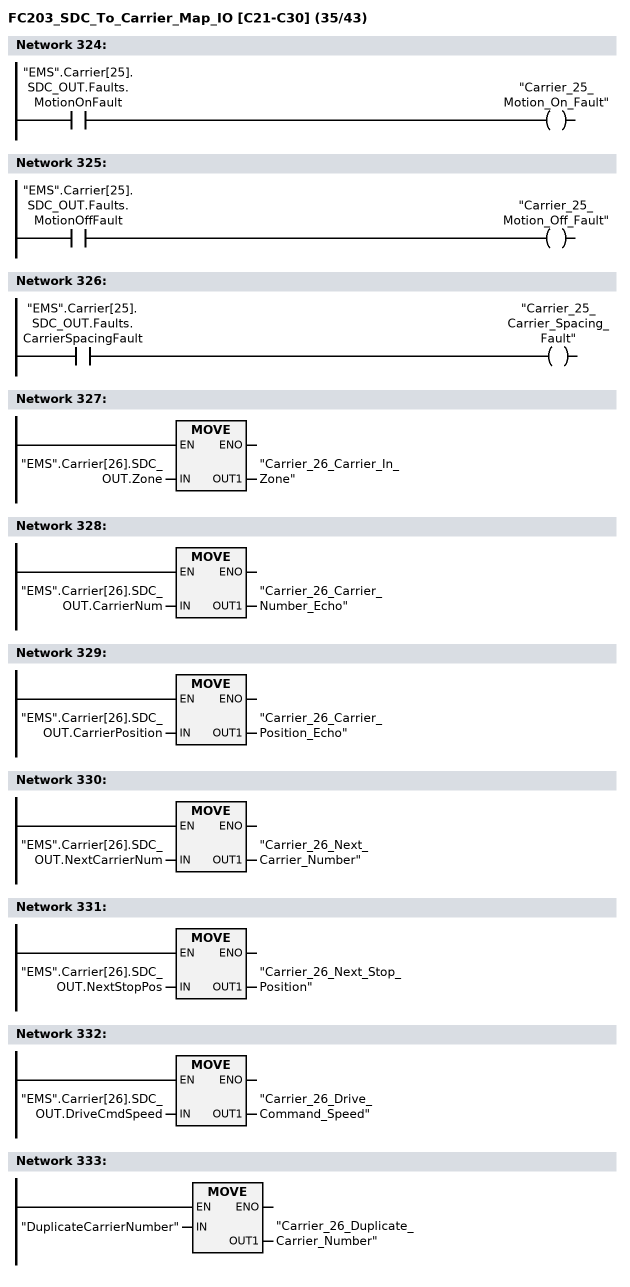
   RUNG wire#powerrail
      Contact( "EMS".Carrier[25].SDC_OUT.Faults.MotionOnFault )
      Coil( "Carrier_25_Motion_On_Fault" )
   END_RUNG
   // the same network as SCL:
   "Carrier_25_Motion_On_Fault" := "EMS".Carrier[25].SDC_OUT.Faults.MotionOnFault;
END_REGION

REGION Network 325
   RUNG wire#powerrail
      Contact( "EMS".Carrier[25].SDC_OUT.Faults.MotionOffFault )
      Coil( "Carrier_25_Motion_Off_Fault" )
   END_RUNG
   // the same network as SCL:
   "Carrier_25_Motion_Off_Fault" := "EMS".Carrier[25].SDC_OUT.Faults.MotionOffFault;
END_REGION

REGION Network 326
   RUNG wire#powerrail
      Contact( "EMS".Carrier[25].SDC_OUT.Faults.CarrierSpacingFault )
      Coil( "Carrier_25_Carrier_Spacing_Fault" )
   END_RUNG
   // the same network as SCL:
   "Carrier_25_Carrier_Spacing_Fault" := "EMS".Carrier[25].SDC_OUT.Faults.CarrierSpacingFault;
END_REGION

REGION Network 327
   RUNG wire#powerrail
      Move(in := "EMS".Carrier[26].SDC_OUT.Zone, out1 => "Carrier_26_Carrier_In_Zone")
   END_RUNG
   // the same network as SCL:
   "Carrier_26_Carrier_In_Zone" := "EMS".Carrier[26].SDC_OUT.Zone;
END_REGION

REGION Network 328
   RUNG wire#powerrail
      Move(in := "EMS".Carrier[26].SDC_OUT.CarrierNum, out1 => "Carrier_26_Carrier_Number_Echo")
   END_RUNG
   // the same network as SCL:
   "Carrier_26_Carrier_Number_Echo" := "EMS".Carrier[26].SDC_OUT.CarrierNum;
END_REGION

REGION Network 329
   RUNG wire#powerrail
      Move(in := "EMS".Carrier[26].SDC_OUT.CarrierPosition, out1 => "Carrier_26_Carrier_Position_Echo")
   END_RUNG
   // the same network as SCL:
   "Carrier_26_Carrier_Position_Echo" := "EMS".Carrier[26].SDC_OUT.CarrierPosition;
END_REGION

REGION Network 330
   RUNG wire#powerrail
      Move(in := "EMS".Carrier[26].SDC_OUT.NextCarrierNum, out1 => "Carrier_26_Next_Carrier_Number")
   END_RUNG
   // the same network as SCL:
   "Carrier_26_Next_Carrier_Number" := "EMS".Carrier[26].SDC_OUT.NextCarrierNum;
END_REGION

REGION Network 331
   RUNG wire#powerrail
      Move(in := "EMS".Carrier[26].SDC_OUT.NextStopPos, out1 => "Carrier_26_Next_Stop_Position")
   END_RUNG
   // the same network as SCL:
   "Carrier_26_Next_Stop_Position" := "EMS".Carrier[26].SDC_OUT.NextStopPos;
END_REGION

REGION Network 332
   RUNG wire#powerrail
      Move(in := "EMS".Carrier[26].SDC_OUT.DriveCmdSpeed, out1 => "Carrier_26_Drive_Command_Speed")
   END_RUNG
   // the same network as SCL:
   "Carrier_26_Drive_Command_Speed" := "EMS".Carrier[26].SDC_OUT.DriveCmdSpeed;
END_REGION

REGION Network 333
   RUNG wire#powerrail
      Move(in := "DuplicateCarrierNumber", out1 => "Carrier_26_Duplicate_Carrier_Number")
   END_RUNG
   // the same network as SCL:
   "Carrier_26_Duplicate_Carrier_Number" := "DuplicateCarrierNumber";
END_REGION

REGION Network 334
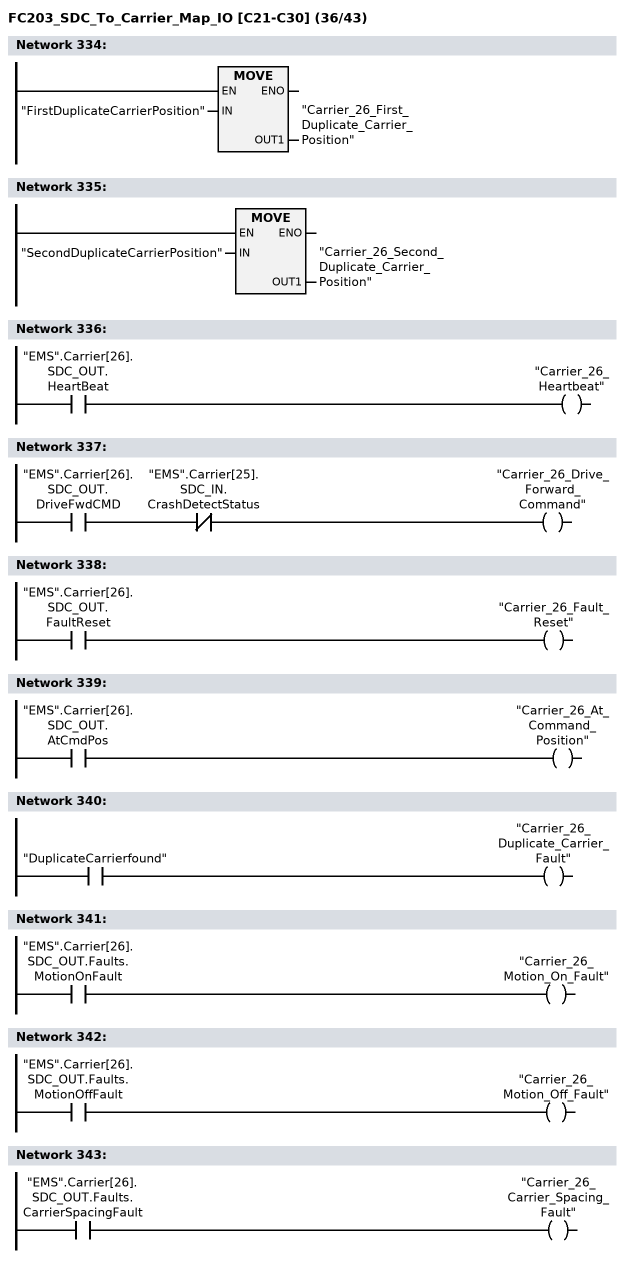
   RUNG wire#powerrail
      Move(in := "FirstDuplicateCarrierPosition", out1 => "Carrier_26_First_Duplicate_Carrier_Position")
   END_RUNG
   // the same network as SCL:
   "Carrier_26_First_Duplicate_Carrier_Position" := "FirstDuplicateCarrierPosition";
END_REGION

REGION Network 335
   RUNG wire#powerrail
      Move(in := "SecondDuplicateCarrierPosition", out1 => "Carrier_26_Second_Duplicate_Carrier_Position")
   END_RUNG
   // the same network as SCL:
   "Carrier_26_Second_Duplicate_Carrier_Position" := "SecondDuplicateCarrierPosition";
END_REGION

REGION Network 336
   RUNG wire#powerrail
      Contact( "EMS".Carrier[26].SDC_OUT.HeartBeat )
      Coil( "Carrier_26_Heartbeat" )
   END_RUNG
   // the same network as SCL:
   "Carrier_26_Heartbeat" := "EMS".Carrier[26].SDC_OUT.HeartBeat;
END_REGION

REGION Network 337
   RUNG wire#powerrail
      Contact( "EMS".Carrier[26].SDC_OUT.DriveFwdCMD )
      I_Contact( "EMS".Carrier[25].SDC_IN.CrashDetectStatus )
      Coil( "Carrier_26_Drive_Forward_Command" )
   END_RUNG
   // the same network as SCL:
   "Carrier_26_Drive_Forward_Command" := "EMS".Carrier[26].SDC_OUT.DriveFwdCMD AND NOT "EMS".Carrier[25].SDC_IN.CrashDetectStatus;
END_REGION

REGION Network 338
   RUNG wire#powerrail
      Contact( "EMS".Carrier[26].SDC_OUT.FaultReset )
      Coil( "Carrier_26_Fault_Reset" )
   END_RUNG
   // the same network as SCL:
   "Carrier_26_Fault_Reset" := "EMS".Carrier[26].SDC_OUT.FaultReset;
END_REGION

REGION Network 339
   RUNG wire#powerrail
      Contact( "EMS".Carrier[26].SDC_OUT.AtCmdPos )
      Coil( "Carrier_26_At_Command_Position" )
   END_RUNG
   // the same network as SCL:
   "Carrier_26_At_Command_Position" := "EMS".Carrier[26].SDC_OUT.AtCmdPos;
END_REGION

REGION Network 340
   RUNG wire#powerrail
      Contact( "DuplicateCarrierfound" )
      Coil( "Carrier_26_Duplicate_Carrier_Fault" )
   END_RUNG
   // the same network as SCL:
   "Carrier_26_Duplicate_Carrier_Fault" := "DuplicateCarrierfound";
END_REGION

REGION Network 341
   RUNG wire#powerrail
      Contact( "EMS".Carrier[26].SDC_OUT.Faults.MotionOnFault )
      Coil( "Carrier_26_Motion_On_Fault" )
   END_RUNG
   // the same network as SCL:
   "Carrier_26_Motion_On_Fault" := "EMS".Carrier[26].SDC_OUT.Faults.MotionOnFault;
END_REGION

REGION Network 342
   RUNG wire#powerrail
      Contact( "EMS".Carrier[26].SDC_OUT.Faults.MotionOffFault )
      Coil( "Carrier_26_Motion_Off_Fault" )
   END_RUNG
   // the same network as SCL:
   "Carrier_26_Motion_Off_Fault" := "EMS".Carrier[26].SDC_OUT.Faults.MotionOffFault;
END_REGION

REGION Network 343
   RUNG wire#powerrail
      Contact( "EMS".Carrier[26].SDC_OUT.Faults.CarrierSpacingFault )
      Coil( "Carrier_26_Carrier_Spacing_Fault" )
   END_RUNG
   // the same network as SCL:
   "Carrier_26_Carrier_Spacing_Fault" := "EMS".Carrier[26].SDC_OUT.Faults.CarrierSpacingFault;
END_REGION

REGION Network 344
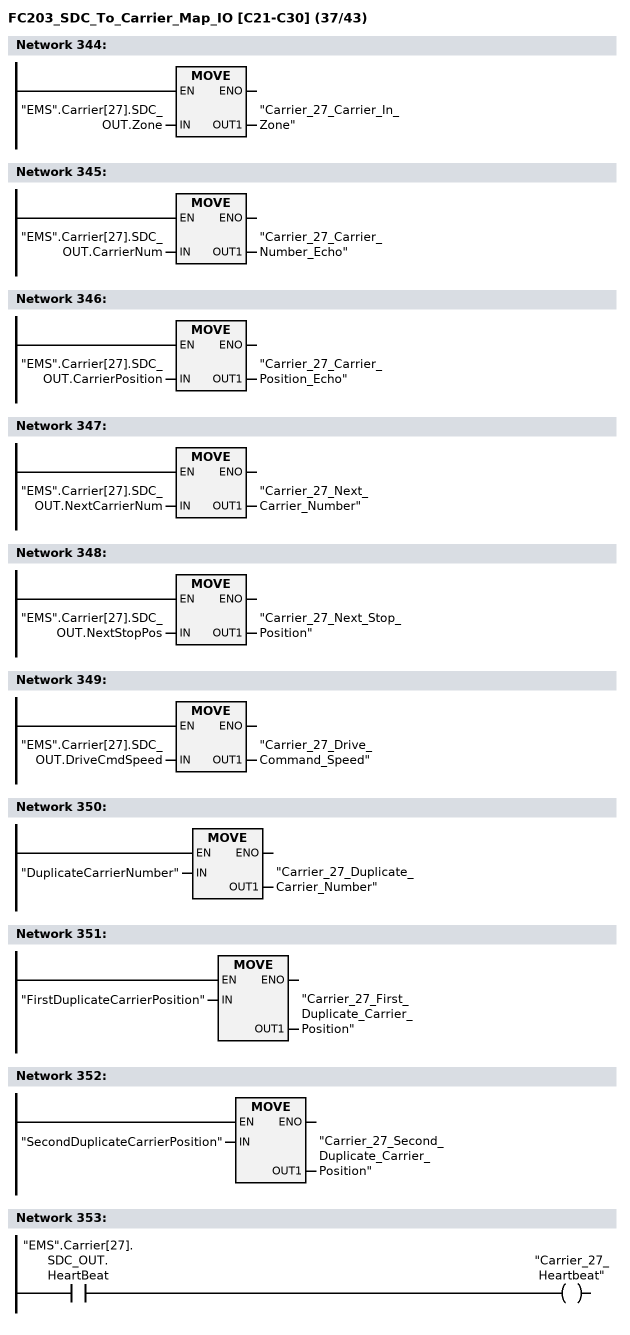
   RUNG wire#powerrail
      Move(in := "EMS".Carrier[27].SDC_OUT.Zone, out1 => "Carrier_27_Carrier_In_Zone")
   END_RUNG
   // the same network as SCL:
   "Carrier_27_Carrier_In_Zone" := "EMS".Carrier[27].SDC_OUT.Zone;
END_REGION

REGION Network 345
   RUNG wire#powerrail
      Move(in := "EMS".Carrier[27].SDC_OUT.CarrierNum, out1 => "Carrier_27_Carrier_Number_Echo")
   END_RUNG
   // the same network as SCL:
   "Carrier_27_Carrier_Number_Echo" := "EMS".Carrier[27].SDC_OUT.CarrierNum;
END_REGION

REGION Network 346
   RUNG wire#powerrail
      Move(in := "EMS".Carrier[27].SDC_OUT.CarrierPosition, out1 => "Carrier_27_Carrier_Position_Echo")
   END_RUNG
   // the same network as SCL:
   "Carrier_27_Carrier_Position_Echo" := "EMS".Carrier[27].SDC_OUT.CarrierPosition;
END_REGION

REGION Network 347
   RUNG wire#powerrail
      Move(in := "EMS".Carrier[27].SDC_OUT.NextCarrierNum, out1 => "Carrier_27_Next_Carrier_Number")
   END_RUNG
   // the same network as SCL:
   "Carrier_27_Next_Carrier_Number" := "EMS".Carrier[27].SDC_OUT.NextCarrierNum;
END_REGION

REGION Network 348
   RUNG wire#powerrail
      Move(in := "EMS".Carrier[27].SDC_OUT.NextStopPos, out1 => "Carrier_27_Next_Stop_Position")
   END_RUNG
   // the same network as SCL:
   "Carrier_27_Next_Stop_Position" := "EMS".Carrier[27].SDC_OUT.NextStopPos;
END_REGION

REGION Network 349
   RUNG wire#powerrail
      Move(in := "EMS".Carrier[27].SDC_OUT.DriveCmdSpeed, out1 => "Carrier_27_Drive_Command_Speed")
   END_RUNG
   // the same network as SCL:
   "Carrier_27_Drive_Command_Speed" := "EMS".Carrier[27].SDC_OUT.DriveCmdSpeed;
END_REGION

REGION Network 350
   RUNG wire#powerrail
      Move(in := "DuplicateCarrierNumber", out1 => "Carrier_27_Duplicate_Carrier_Number")
   END_RUNG
   // the same network as SCL:
   "Carrier_27_Duplicate_Carrier_Number" := "DuplicateCarrierNumber";
END_REGION

REGION Network 351
   RUNG wire#powerrail
      Move(in := "FirstDuplicateCarrierPosition", out1 => "Carrier_27_First_Duplicate_Carrier_Position")
   END_RUNG
   // the same network as SCL:
   "Carrier_27_First_Duplicate_Carrier_Position" := "FirstDuplicateCarrierPosition";
END_REGION

REGION Network 352
   RUNG wire#powerrail
      Move(in := "SecondDuplicateCarrierPosition", out1 => "Carrier_27_Second_Duplicate_Carrier_Position")
   END_RUNG
   // the same network as SCL:
   "Carrier_27_Second_Duplicate_Carrier_Position" := "SecondDuplicateCarrierPosition";
END_REGION

REGION Network 353
   RUNG wire#powerrail
      Contact( "EMS".Carrier[27].SDC_OUT.HeartBeat )
      Coil( "Carrier_27_Heartbeat" )
   END_RUNG
   // the same network as SCL:
   "Carrier_27_Heartbeat" := "EMS".Carrier[27].SDC_OUT.HeartBeat;
END_REGION

REGION Network 354
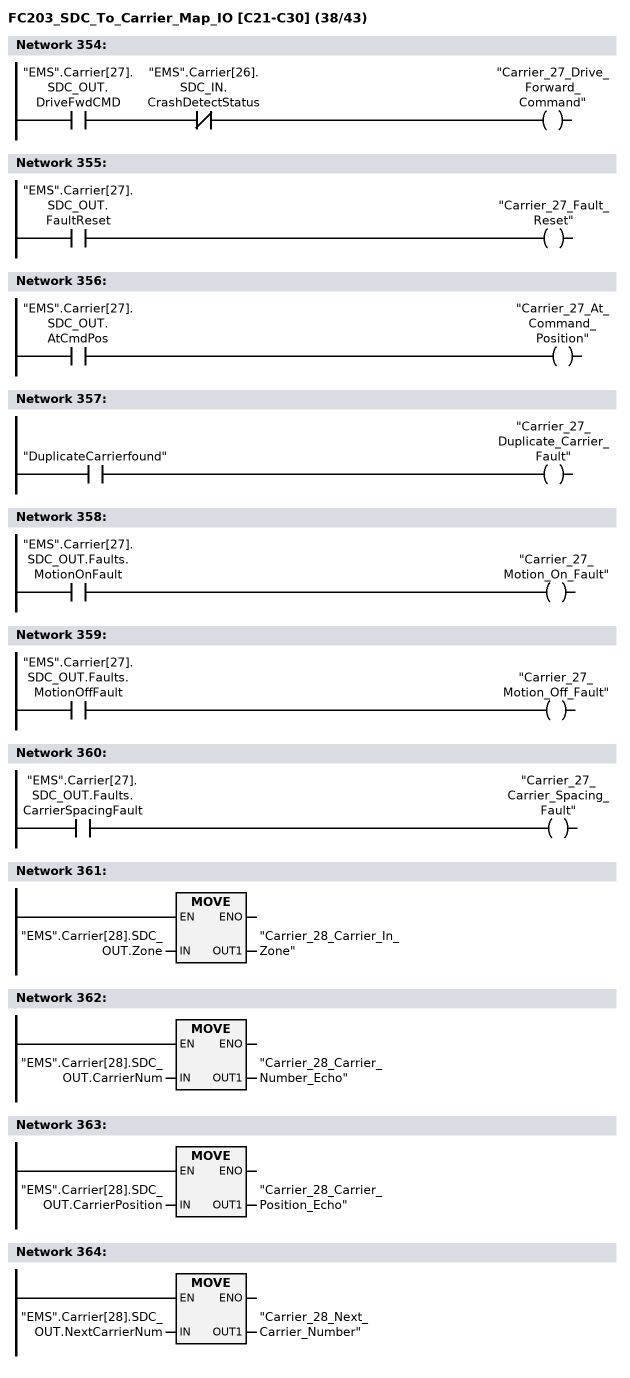
   RUNG wire#powerrail
      Contact( "EMS".Carrier[27].SDC_OUT.DriveFwdCMD )
      I_Contact( "EMS".Carrier[26].SDC_IN.CrashDetectStatus )
      Coil( "Carrier_27_Drive_Forward_Command" )
   END_RUNG
   // the same network as SCL:
   "Carrier_27_Drive_Forward_Command" := "EMS".Carrier[27].SDC_OUT.DriveFwdCMD AND NOT "EMS".Carrier[26].SDC_IN.CrashDetectStatus;
END_REGION

REGION Network 355
   RUNG wire#powerrail
      Contact( "EMS".Carrier[27].SDC_OUT.FaultReset )
      Coil( "Carrier_27_Fault_Reset" )
   END_RUNG
   // the same network as SCL:
   "Carrier_27_Fault_Reset" := "EMS".Carrier[27].SDC_OUT.FaultReset;
END_REGION

REGION Network 356
   RUNG wire#powerrail
      Contact( "EMS".Carrier[27].SDC_OUT.AtCmdPos )
      Coil( "Carrier_27_At_Command_Position" )
   END_RUNG
   // the same network as SCL:
   "Carrier_27_At_Command_Position" := "EMS".Carrier[27].SDC_OUT.AtCmdPos;
END_REGION

REGION Network 357
   RUNG wire#powerrail
      Contact( "DuplicateCarrierfound" )
      Coil( "Carrier_27_Duplicate_Carrier_Fault" )
   END_RUNG
   // the same network as SCL:
   "Carrier_27_Duplicate_Carrier_Fault" := "DuplicateCarrierfound";
END_REGION

REGION Network 358
   RUNG wire#powerrail
      Contact( "EMS".Carrier[27].SDC_OUT.Faults.MotionOnFault )
      Coil( "Carrier_27_Motion_On_Fault" )
   END_RUNG
   // the same network as SCL:
   "Carrier_27_Motion_On_Fault" := "EMS".Carrier[27].SDC_OUT.Faults.MotionOnFault;
END_REGION

REGION Network 359
   RUNG wire#powerrail
      Contact( "EMS".Carrier[27].SDC_OUT.Faults.MotionOffFault )
      Coil( "Carrier_27_Motion_Off_Fault" )
   END_RUNG
   // the same network as SCL:
   "Carrier_27_Motion_Off_Fault" := "EMS".Carrier[27].SDC_OUT.Faults.MotionOffFault;
END_REGION

REGION Network 360
   RUNG wire#powerrail
      Contact( "EMS".Carrier[27].SDC_OUT.Faults.CarrierSpacingFault )
      Coil( "Carrier_27_Carrier_Spacing_Fault" )
   END_RUNG
   // the same network as SCL:
   "Carrier_27_Carrier_Spacing_Fault" := "EMS".Carrier[27].SDC_OUT.Faults.CarrierSpacingFault;
END_REGION

REGION Network 361
   RUNG wire#powerrail
      Move(in := "EMS".Carrier[28].SDC_OUT.Zone, out1 => "Carrier_28_Carrier_In_Zone")
   END_RUNG
   // the same network as SCL:
   "Carrier_28_Carrier_In_Zone" := "EMS".Carrier[28].SDC_OUT.Zone;
END_REGION

REGION Network 362
   RUNG wire#powerrail
      Move(in := "EMS".Carrier[28].SDC_OUT.CarrierNum, out1 => "Carrier_28_Carrier_Number_Echo")
   END_RUNG
   // the same network as SCL:
   "Carrier_28_Carrier_Number_Echo" := "EMS".Carrier[28].SDC_OUT.CarrierNum;
END_REGION

REGION Network 363
   RUNG wire#powerrail
      Move(in := "EMS".Carrier[28].SDC_OUT.CarrierPosition, out1 => "Carrier_28_Carrier_Position_Echo")
   END_RUNG
   // the same network as SCL:
   "Carrier_28_Carrier_Position_Echo" := "EMS".Carrier[28].SDC_OUT.CarrierPosition;
END_REGION

REGION Network 364
   RUNG wire#powerrail
      Move(in := "EMS".Carrier[28].SDC_OUT.NextCarrierNum, out1 => "Carrier_28_Next_Carrier_Number")
   END_RUNG
   // the same network as SCL:
   "Carrier_28_Next_Carrier_Number" := "EMS".Carrier[28].SDC_OUT.NextCarrierNum;
END_REGION

REGION Network 365
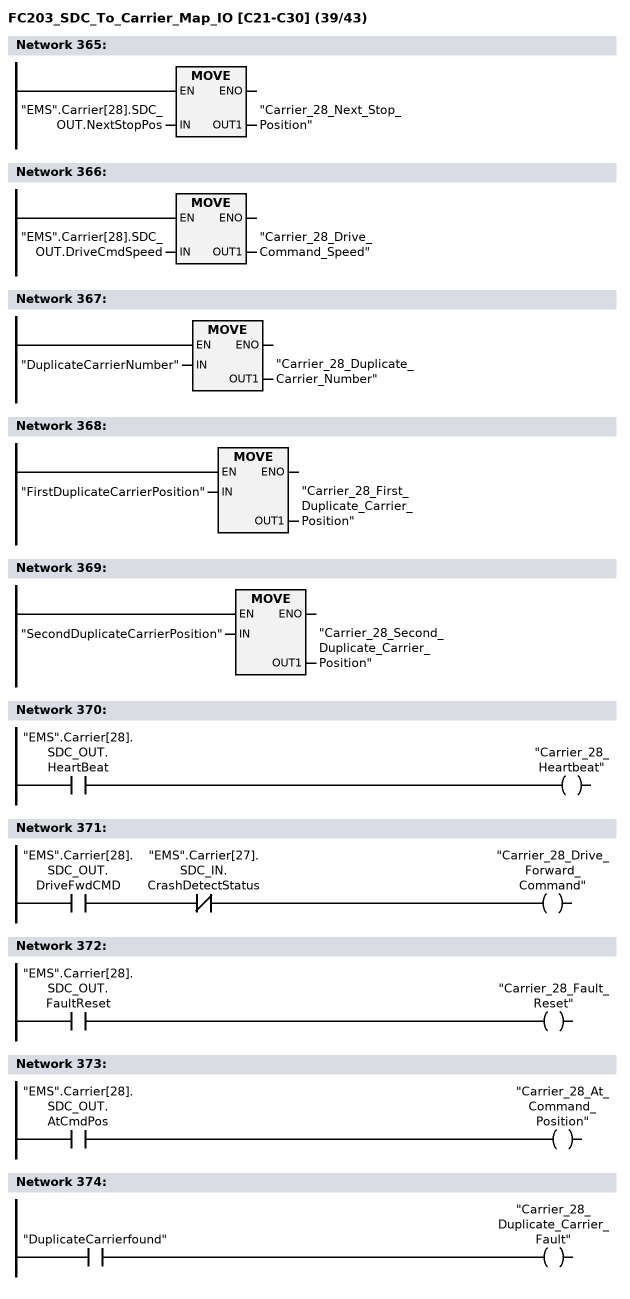
   RUNG wire#powerrail
      Move(in := "EMS".Carrier[28].SDC_OUT.NextStopPos, out1 => "Carrier_28_Next_Stop_Position")
   END_RUNG
   // the same network as SCL:
   "Carrier_28_Next_Stop_Position" := "EMS".Carrier[28].SDC_OUT.NextStopPos;
END_REGION

REGION Network 366
   RUNG wire#powerrail
      Move(in := "EMS".Carrier[28].SDC_OUT.DriveCmdSpeed, out1 => "Carrier_28_Drive_Command_Speed")
   END_RUNG
   // the same network as SCL:
   "Carrier_28_Drive_Command_Speed" := "EMS".Carrier[28].SDC_OUT.DriveCmdSpeed;
END_REGION

REGION Network 367
   RUNG wire#powerrail
      Move(in := "DuplicateCarrierNumber", out1 => "Carrier_28_Duplicate_Carrier_Number")
   END_RUNG
   // the same network as SCL:
   "Carrier_28_Duplicate_Carrier_Number" := "DuplicateCarrierNumber";
END_REGION

REGION Network 368
   RUNG wire#powerrail
      Move(in := "FirstDuplicateCarrierPosition", out1 => "Carrier_28_First_Duplicate_Carrier_Position")
   END_RUNG
   // the same network as SCL:
   "Carrier_28_First_Duplicate_Carrier_Position" := "FirstDuplicateCarrierPosition";
END_REGION

REGION Network 369
   RUNG wire#powerrail
      Move(in := "SecondDuplicateCarrierPosition", out1 => "Carrier_28_Second_Duplicate_Carrier_Position")
   END_RUNG
   // the same network as SCL:
   "Carrier_28_Second_Duplicate_Carrier_Position" := "SecondDuplicateCarrierPosition";
END_REGION

REGION Network 370
   RUNG wire#powerrail
      Contact( "EMS".Carrier[28].SDC_OUT.HeartBeat )
      Coil( "Carrier_28_Heartbeat" )
   END_RUNG
   // the same network as SCL:
   "Carrier_28_Heartbeat" := "EMS".Carrier[28].SDC_OUT.HeartBeat;
END_REGION

REGION Network 371
   RUNG wire#powerrail
      Contact( "EMS".Carrier[28].SDC_OUT.DriveFwdCMD )
      I_Contact( "EMS".Carrier[27].SDC_IN.CrashDetectStatus )
      Coil( "Carrier_28_Drive_Forward_Command" )
   END_RUNG
   // the same network as SCL:
   "Carrier_28_Drive_Forward_Command" := "EMS".Carrier[28].SDC_OUT.DriveFwdCMD AND NOT "EMS".Carrier[27].SDC_IN.CrashDetectStatus;
END_REGION

REGION Network 372
   RUNG wire#powerrail
      Contact( "EMS".Carrier[28].SDC_OUT.FaultReset )
      Coil( "Carrier_28_Fault_Reset" )
   END_RUNG
   // the same network as SCL:
   "Carrier_28_Fault_Reset" := "EMS".Carrier[28].SDC_OUT.FaultReset;
END_REGION

REGION Network 373
   RUNG wire#powerrail
      Contact( "EMS".Carrier[28].SDC_OUT.AtCmdPos )
      Coil( "Carrier_28_At_Command_Position" )
   END_RUNG
   // the same network as SCL:
   "Carrier_28_At_Command_Position" := "EMS".Carrier[28].SDC_OUT.AtCmdPos;
END_REGION

REGION Network 374
   RUNG wire#powerrail
      Contact( "DuplicateCarrierfound" )
      Coil( "Carrier_28_Duplicate_Carrier_Fault" )
   END_RUNG
   // the same network as SCL:
   "Carrier_28_Duplicate_Carrier_Fault" := "DuplicateCarrierfound";
END_REGION

REGION Network 375
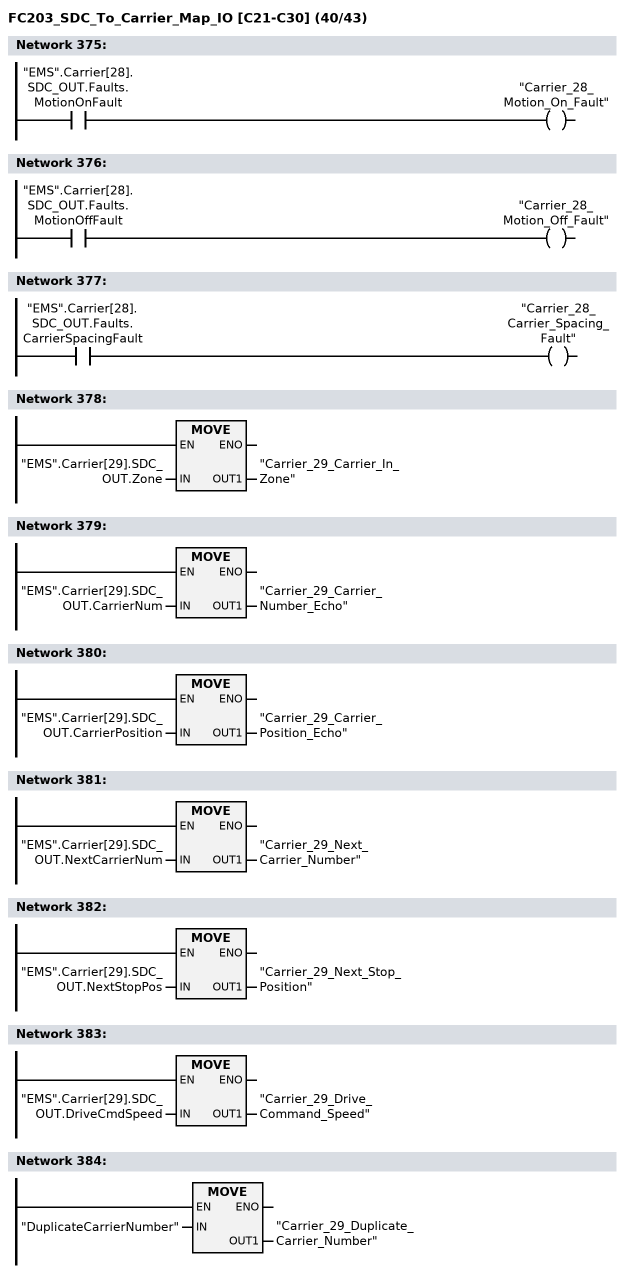
   RUNG wire#powerrail
      Contact( "EMS".Carrier[28].SDC_OUT.Faults.MotionOnFault )
      Coil( "Carrier_28_Motion_On_Fault" )
   END_RUNG
   // the same network as SCL:
   "Carrier_28_Motion_On_Fault" := "EMS".Carrier[28].SDC_OUT.Faults.MotionOnFault;
END_REGION

REGION Network 376
   RUNG wire#powerrail
      Contact( "EMS".Carrier[28].SDC_OUT.Faults.MotionOffFault )
      Coil( "Carrier_28_Motion_Off_Fault" )
   END_RUNG
   // the same network as SCL:
   "Carrier_28_Motion_Off_Fault" := "EMS".Carrier[28].SDC_OUT.Faults.MotionOffFault;
END_REGION

REGION Network 377
   RUNG wire#powerrail
      Contact( "EMS".Carrier[28].SDC_OUT.Faults.CarrierSpacingFault )
      Coil( "Carrier_28_Carrier_Spacing_Fault" )
   END_RUNG
   // the same network as SCL:
   "Carrier_28_Carrier_Spacing_Fault" := "EMS".Carrier[28].SDC_OUT.Faults.CarrierSpacingFault;
END_REGION

REGION Network 378
   RUNG wire#powerrail
      Move(in := "EMS".Carrier[29].SDC_OUT.Zone, out1 => "Carrier_29_Carrier_In_Zone")
   END_RUNG
   // the same network as SCL:
   "Carrier_29_Carrier_In_Zone" := "EMS".Carrier[29].SDC_OUT.Zone;
END_REGION

REGION Network 379
   RUNG wire#powerrail
      Move(in := "EMS".Carrier[29].SDC_OUT.CarrierNum, out1 => "Carrier_29_Carrier_Number_Echo")
   END_RUNG
   // the same network as SCL:
   "Carrier_29_Carrier_Number_Echo" := "EMS".Carrier[29].SDC_OUT.CarrierNum;
END_REGION

REGION Network 380
   RUNG wire#powerrail
      Move(in := "EMS".Carrier[29].SDC_OUT.CarrierPosition, out1 => "Carrier_29_Carrier_Position_Echo")
   END_RUNG
   // the same network as SCL:
   "Carrier_29_Carrier_Position_Echo" := "EMS".Carrier[29].SDC_OUT.CarrierPosition;
END_REGION

REGION Network 381
   RUNG wire#powerrail
      Move(in := "EMS".Carrier[29].SDC_OUT.NextCarrierNum, out1 => "Carrier_29_Next_Carrier_Number")
   END_RUNG
   // the same network as SCL:
   "Carrier_29_Next_Carrier_Number" := "EMS".Carrier[29].SDC_OUT.NextCarrierNum;
END_REGION

REGION Network 382
   RUNG wire#powerrail
      Move(in := "EMS".Carrier[29].SDC_OUT.NextStopPos, out1 => "Carrier_29_Next_Stop_Position")
   END_RUNG
   // the same network as SCL:
   "Carrier_29_Next_Stop_Position" := "EMS".Carrier[29].SDC_OUT.NextStopPos;
END_REGION

REGION Network 383
   RUNG wire#powerrail
      Move(in := "EMS".Carrier[29].SDC_OUT.DriveCmdSpeed, out1 => "Carrier_29_Drive_Command_Speed")
   END_RUNG
   // the same network as SCL:
   "Carrier_29_Drive_Command_Speed" := "EMS".Carrier[29].SDC_OUT.DriveCmdSpeed;
END_REGION

REGION Network 384
   RUNG wire#powerrail
      Move(in := "DuplicateCarrierNumber", out1 => "Carrier_29_Duplicate_Carrier_Number")
   END_RUNG
   // the same network as SCL:
   "Carrier_29_Duplicate_Carrier_Number" := "DuplicateCarrierNumber";
END_REGION

REGION Network 385
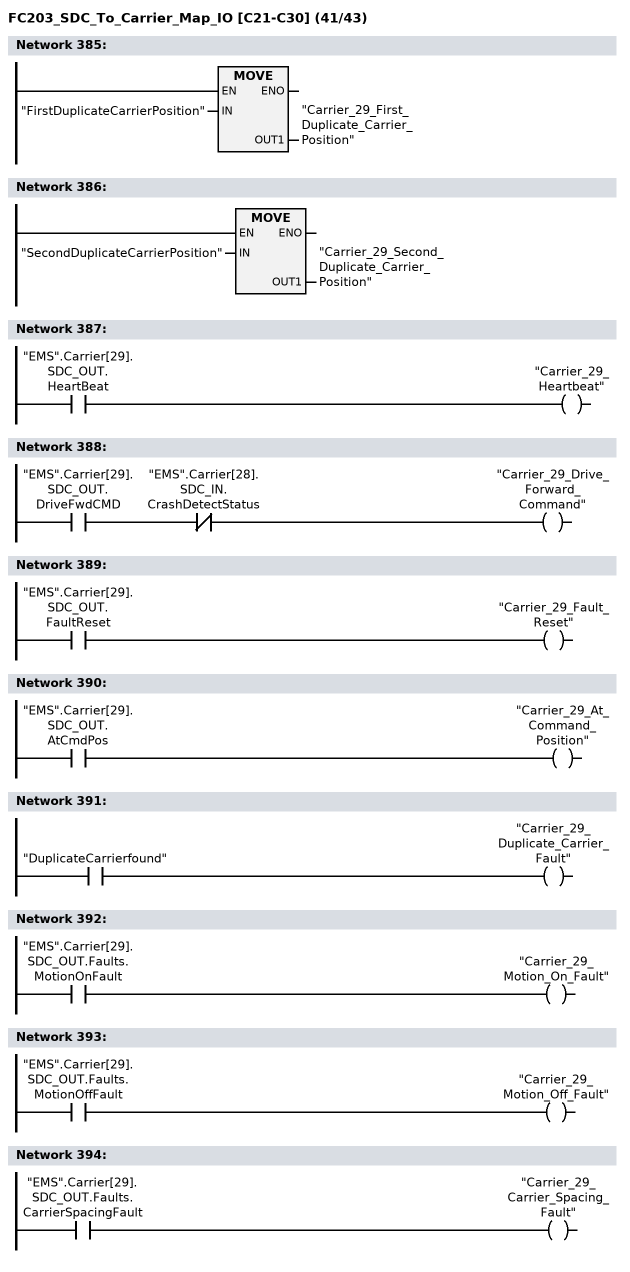
   RUNG wire#powerrail
      Move(in := "FirstDuplicateCarrierPosition", out1 => "Carrier_29_First_Duplicate_Carrier_Position")
   END_RUNG
   // the same network as SCL:
   "Carrier_29_First_Duplicate_Carrier_Position" := "FirstDuplicateCarrierPosition";
END_REGION

REGION Network 386
   RUNG wire#powerrail
      Move(in := "SecondDuplicateCarrierPosition", out1 => "Carrier_29_Second_Duplicate_Carrier_Position")
   END_RUNG
   // the same network as SCL:
   "Carrier_29_Second_Duplicate_Carrier_Position" := "SecondDuplicateCarrierPosition";
END_REGION

REGION Network 387
   RUNG wire#powerrail
      Contact( "EMS".Carrier[29].SDC_OUT.HeartBeat )
      Coil( "Carrier_29_Heartbeat" )
   END_RUNG
   // the same network as SCL:
   "Carrier_29_Heartbeat" := "EMS".Carrier[29].SDC_OUT.HeartBeat;
END_REGION

REGION Network 388
   RUNG wire#powerrail
      Contact( "EMS".Carrier[29].SDC_OUT.DriveFwdCMD )
      I_Contact( "EMS".Carrier[28].SDC_IN.CrashDetectStatus )
      Coil( "Carrier_29_Drive_Forward_Command" )
   END_RUNG
   // the same network as SCL:
   "Carrier_29_Drive_Forward_Command" := "EMS".Carrier[29].SDC_OUT.DriveFwdCMD AND NOT "EMS".Carrier[28].SDC_IN.CrashDetectStatus;
END_REGION

REGION Network 389
   RUNG wire#powerrail
      Contact( "EMS".Carrier[29].SDC_OUT.FaultReset )
      Coil( "Carrier_29_Fault_Reset" )
   END_RUNG
   // the same network as SCL:
   "Carrier_29_Fault_Reset" := "EMS".Carrier[29].SDC_OUT.FaultReset;
END_REGION

REGION Network 390
   RUNG wire#powerrail
      Contact( "EMS".Carrier[29].SDC_OUT.AtCmdPos )
      Coil( "Carrier_29_At_Command_Position" )
   END_RUNG
   // the same network as SCL:
   "Carrier_29_At_Command_Position" := "EMS".Carrier[29].SDC_OUT.AtCmdPos;
END_REGION

REGION Network 391
   RUNG wire#powerrail
      Contact( "DuplicateCarrierfound" )
      Coil( "Carrier_29_Duplicate_Carrier_Fault" )
   END_RUNG
   // the same network as SCL:
   "Carrier_29_Duplicate_Carrier_Fault" := "DuplicateCarrierfound";
END_REGION

REGION Network 392
   RUNG wire#powerrail
      Contact( "EMS".Carrier[29].SDC_OUT.Faults.MotionOnFault )
      Coil( "Carrier_29_Motion_On_Fault" )
   END_RUNG
   // the same network as SCL:
   "Carrier_29_Motion_On_Fault" := "EMS".Carrier[29].SDC_OUT.Faults.MotionOnFault;
END_REGION

REGION Network 393
   RUNG wire#powerrail
      Contact( "EMS".Carrier[29].SDC_OUT.Faults.MotionOffFault )
      Coil( "Carrier_29_Motion_Off_Fault" )
   END_RUNG
   // the same network as SCL:
   "Carrier_29_Motion_Off_Fault" := "EMS".Carrier[29].SDC_OUT.Faults.MotionOffFault;
END_REGION

REGION Network 394
   RUNG wire#powerrail
      Contact( "EMS".Carrier[29].SDC_OUT.Faults.CarrierSpacingFault )
      Coil( "Carrier_29_Carrier_Spacing_Fault" )
   END_RUNG
   // the same network as SCL:
   "Carrier_29_Carrier_Spacing_Fault" := "EMS".Carrier[29].SDC_OUT.Faults.CarrierSpacingFault;
END_REGION

REGION Network 395
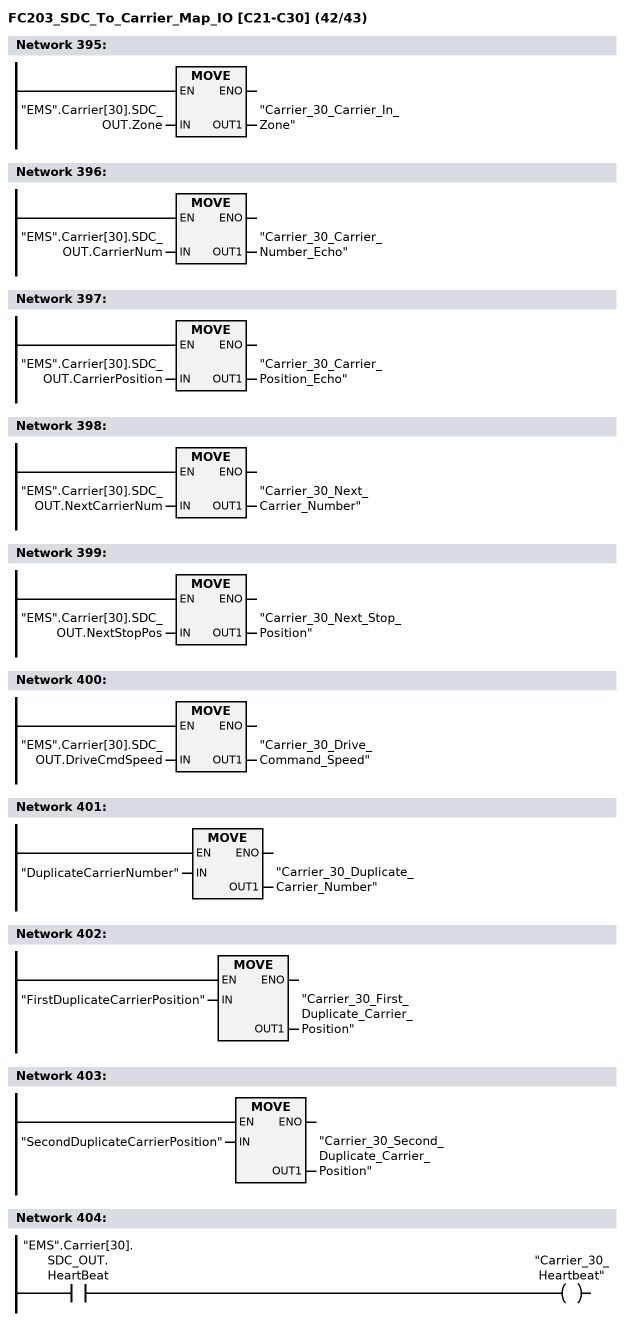
   RUNG wire#powerrail
      Move(in := "EMS".Carrier[30].SDC_OUT.Zone, out1 => "Carrier_30_Carrier_In_Zone")
   END_RUNG
   // the same network as SCL:
   "Carrier_30_Carrier_In_Zone" := "EMS".Carrier[30].SDC_OUT.Zone;
END_REGION

REGION Network 396
   RUNG wire#powerrail
      Move(in := "EMS".Carrier[30].SDC_OUT.CarrierNum, out1 => "Carrier_30_Carrier_Number_Echo")
   END_RUNG
   // the same network as SCL:
   "Carrier_30_Carrier_Number_Echo" := "EMS".Carrier[30].SDC_OUT.CarrierNum;
END_REGION

REGION Network 397
   RUNG wire#powerrail
      Move(in := "EMS".Carrier[30].SDC_OUT.CarrierPosition, out1 => "Carrier_30_Carrier_Position_Echo")
   END_RUNG
   // the same network as SCL:
   "Carrier_30_Carrier_Position_Echo" := "EMS".Carrier[30].SDC_OUT.CarrierPosition;
END_REGION

REGION Network 398
   RUNG wire#powerrail
      Move(in := "EMS".Carrier[30].SDC_OUT.NextCarrierNum, out1 => "Carrier_30_Next_Carrier_Number")
   END_RUNG
   // the same network as SCL:
   "Carrier_30_Next_Carrier_Number" := "EMS".Carrier[30].SDC_OUT.NextCarrierNum;
END_REGION

REGION Network 399
   RUNG wire#powerrail
      Move(in := "EMS".Carrier[30].SDC_OUT.NextStopPos, out1 => "Carrier_30_Next_Stop_Position")
   END_RUNG
   // the same network as SCL:
   "Carrier_30_Next_Stop_Position" := "EMS".Carrier[30].SDC_OUT.NextStopPos;
END_REGION

REGION Network 400
   RUNG wire#powerrail
      Move(in := "EMS".Carrier[30].SDC_OUT.DriveCmdSpeed, out1 => "Carrier_30_Drive_Command_Speed")
   END_RUNG
   // the same network as SCL:
   "Carrier_30_Drive_Command_Speed" := "EMS".Carrier[30].SDC_OUT.DriveCmdSpeed;
END_REGION

REGION Network 401
   RUNG wire#powerrail
      Move(in := "DuplicateCarrierNumber", out1 => "Carrier_30_Duplicate_Carrier_Number")
   END_RUNG
   // the same network as SCL:
   "Carrier_30_Duplicate_Carrier_Number" := "DuplicateCarrierNumber";
END_REGION

REGION Network 402
   RUNG wire#powerrail
      Move(in := "FirstDuplicateCarrierPosition", out1 => "Carrier_30_First_Duplicate_Carrier_Position")
   END_RUNG
   // the same network as SCL:
   "Carrier_30_First_Duplicate_Carrier_Position" := "FirstDuplicateCarrierPosition";
END_REGION

REGION Network 403
   RUNG wire#powerrail
      Move(in := "SecondDuplicateCarrierPosition", out1 => "Carrier_30_Second_Duplicate_Carrier_Position")
   END_RUNG
   // the same network as SCL:
   "Carrier_30_Second_Duplicate_Carrier_Position" := "SecondDuplicateCarrierPosition";
END_REGION

REGION Network 404
   RUNG wire#powerrail
      Contact( "EMS".Carrier[30].SDC_OUT.HeartBeat )
      Coil( "Carrier_30_Heartbeat" )
   END_RUNG
   // the same network as SCL:
   "Carrier_30_Heartbeat" := "EMS".Carrier[30].SDC_OUT.HeartBeat;
END_REGION

REGION Network 405
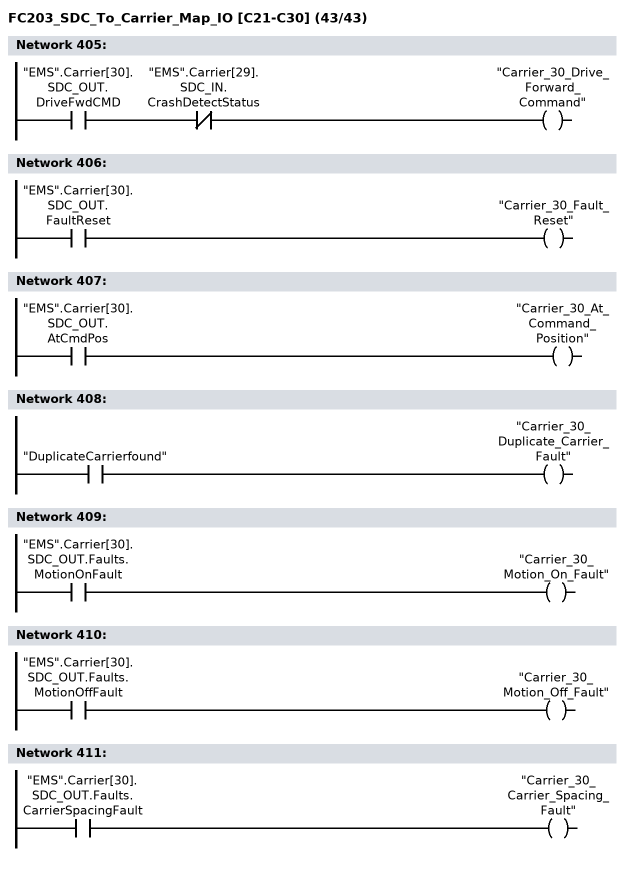
   RUNG wire#powerrail
      Contact( "EMS".Carrier[30].SDC_OUT.DriveFwdCMD )
      I_Contact( "EMS".Carrier[29].SDC_IN.CrashDetectStatus )
      Coil( "Carrier_30_Drive_Forward_Command" )
   END_RUNG
   // the same network as SCL:
   "Carrier_30_Drive_Forward_Command" := "EMS".Carrier[30].SDC_OUT.DriveFwdCMD AND NOT "EMS".Carrier[29].SDC_IN.CrashDetectStatus;
END_REGION

REGION Network 406
   RUNG wire#powerrail
      Contact( "EMS".Carrier[30].SDC_OUT.FaultReset )
      Coil( "Carrier_30_Fault_Reset" )
   END_RUNG
   // the same network as SCL:
   "Carrier_30_Fault_Reset" := "EMS".Carrier[30].SDC_OUT.FaultReset;
END_REGION

REGION Network 407
   RUNG wire#powerrail
      Contact( "EMS".Carrier[30].SDC_OUT.AtCmdPos )
      Coil( "Carrier_30_At_Command_Position" )
   END_RUNG
   // the same network as SCL:
   "Carrier_30_At_Command_Position" := "EMS".Carrier[30].SDC_OUT.AtCmdPos;
END_REGION

REGION Network 408
   RUNG wire#powerrail
      Contact( "DuplicateCarrierfound" )
      Coil( "Carrier_30_Duplicate_Carrier_Fault" )
   END_RUNG
   // the same network as SCL:
   "Carrier_30_Duplicate_Carrier_Fault" := "DuplicateCarrierfound";
END_REGION

REGION Network 409
   RUNG wire#powerrail
      Contact( "EMS".Carrier[30].SDC_OUT.Faults.MotionOnFault )
      Coil( "Carrier_30_Motion_On_Fault" )
   END_RUNG
   // the same network as SCL:
   "Carrier_30_Motion_On_Fault" := "EMS".Carrier[30].SDC_OUT.Faults.MotionOnFault;
END_REGION

REGION Network 410
   RUNG wire#powerrail
      Contact( "EMS".Carrier[30].SDC_OUT.Faults.MotionOffFault )
      Coil( "Carrier_30_Motion_Off_Fault" )
   END_RUNG
   // the same network as SCL:
   "Carrier_30_Motion_Off_Fault" := "EMS".Carrier[30].SDC_OUT.Faults.MotionOffFault;
END_REGION

REGION Network 411
   RUNG wire#powerrail
      Contact( "EMS".Carrier[30].SDC_OUT.Faults.CarrierSpacingFault )
      Coil( "Carrier_30_Carrier_Spacing_Fault" )
   END_RUNG
   // the same network as SCL:
   "Carrier_30_Carrier_Spacing_Fault" := "EMS".Carrier[30].SDC_OUT.Faults.CarrierSpacingFault;
END_REGION
END_FUNCTION

FUNCTION "FC204_SDC_To_Carrier_Map_IO [C31-C40]" : Void   // FC204, LAD
{ S7_Optimized_Access := 'TRUE' }
VERSION : 0.1
BEGIN

REGION Network 1